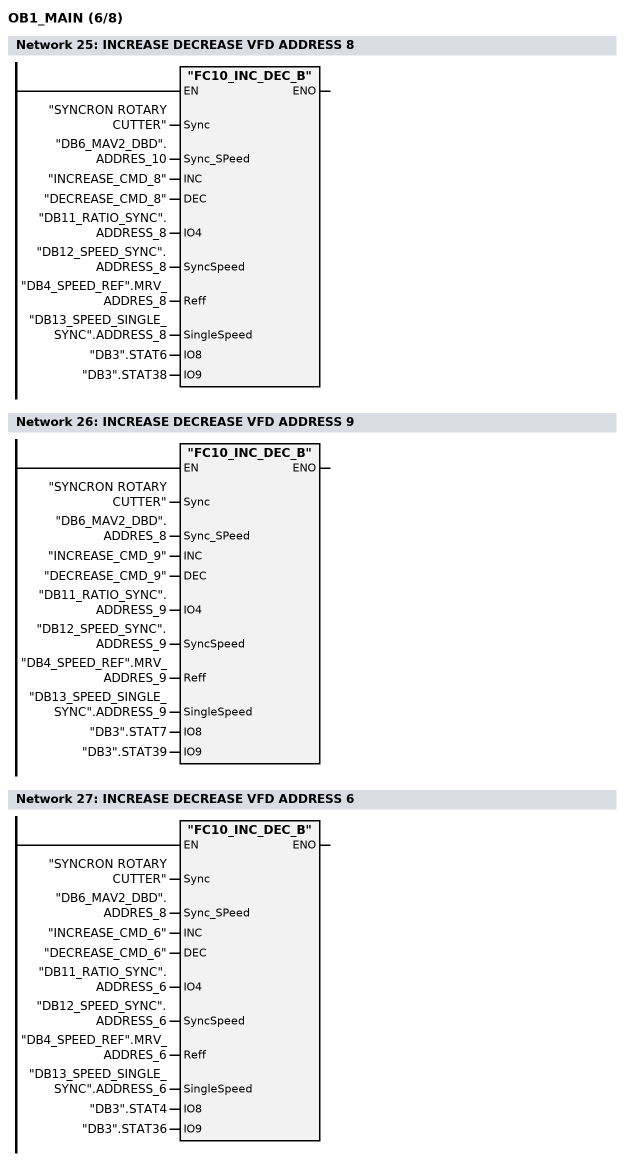
   RUNG wire#powerrail
      "FC10_INC_DEC_B"(Sync := "SYNCRON ROTARY CUTTER", Sync_SPeed := "DB6_MAV2_DBD".ADDRES_10, INC := "INCREASE_CMD_8", DEC := "DECREASE_CMD_8", IO4 := "DB11_RATIO_SYNC".ADDRESS_8, SyncSpeed := "DB12_SPEED_SYNC".ADDRESS_8, Reff := "DB4_SPEED_REF".MRV_ADDRES_8, SingleSpeed := "DB13_SPEED_SINGLE_SYNC".ADDRESS_8, IO8 := "DB3".STAT6, IO9 := "DB3".STAT38)
   END_RUNG
   // the same network as SCL:
   "FC10_INC_DEC_B"(Sync := "SYNCRON ROTARY CUTTER",
                    Sync_SPeed := "DB6_MAV2_DBD".ADDRES_10,
                    INC := "INCREASE_CMD_8",
                    DEC := "DECREASE_CMD_8",
                    IO4 := "DB11_RATIO_SYNC".ADDRESS_8,
                    SyncSpeed := "DB12_SPEED_SYNC".ADDRESS_8,
                    Reff := "DB4_SPEED_REF".MRV_ADDRES_8,
                    SingleSpeed := "DB13_SPEED_SINGLE_SYNC".ADDRESS_8,
                    IO8 := "DB3".STAT6,
                    IO9 := "DB3".STAT38);
END_REGION

REGION Network 26: INCREASE DECREASE VFD ADDRESS 9
   RUNG wire#powerrail
      "FC10_INC_DEC_B"(Sync := "SYNCRON ROTARY CUTTER", Sync_SPeed := "DB6_MAV2_DBD".ADDRES_8, INC := "INCREASE_CMD_9", DEC := "DECREASE_CMD_9", IO4 := "DB11_RATIO_SYNC".ADDRESS_9, SyncSpeed := "DB12_SPEED_SYNC".ADDRESS_9, Reff := "DB4_SPEED_REF".MRV_ADDRES_9, SingleSpeed := "DB13_SPEED_SINGLE_SYNC".ADDRESS_9, IO8 := "DB3".STAT7, IO9 := "DB3".STAT39)
   END_RUNG
   // the same network as SCL:
   "FC10_INC_DEC_B"(Sync := "SYNCRON ROTARY CUTTER",
                    Sync_SPeed := "DB6_MAV2_DBD".ADDRES_8,
                    INC := "INCREASE_CMD_9",
                    DEC := "DECREASE_CMD_9",
                    IO4 := "DB11_RATIO_SYNC".ADDRESS_9,
                    SyncSpeed := "DB12_SPEED_SYNC".ADDRESS_9,
                    Reff := "DB4_SPEED_REF".MRV_ADDRES_9,
                    SingleSpeed := "DB13_SPEED_SINGLE_SYNC".ADDRESS_9,
                    IO8 := "DB3".STAT7,
                    IO9 := "DB3".STAT39);
END_REGION

REGION Network 27: INCREASE DECREASE VFD ADDRESS 6
   RUNG wire#powerrail
      "FC10_INC_DEC_B"(Sync := "SYNCRON ROTARY CUTTER", Sync_SPeed := "DB6_MAV2_DBD".ADDRES_8, INC := "INCREASE_CMD_6", DEC := "DECREASE_CMD_6", IO4 := "DB11_RATIO_SYNC".ADDRESS_6, SyncSpeed := "DB12_SPEED_SYNC".ADDRESS_6, Reff := "DB4_SPEED_REF".MRV_ADDRES_6, SingleSpeed := "DB13_SPEED_SINGLE_SYNC".ADDRESS_6, IO8 := "DB3".STAT4, IO9 := "DB3".STAT36)
   END_RUNG
   // the same network as SCL:
   "FC10_INC_DEC_B"(Sync := "SYNCRON ROTARY CUTTER",
                    Sync_SPeed := "DB6_MAV2_DBD".ADDRES_8,
                    INC := "INCREASE_CMD_6",
                    DEC := "DECREASE_CMD_6",
                    IO4 := "DB11_RATIO_SYNC".ADDRESS_6,
                    SyncSpeed := "DB12_SPEED_SYNC".ADDRESS_6,
                    Reff := "DB4_SPEED_REF".MRV_ADDRES_6,
                    SingleSpeed := "DB13_SPEED_SINGLE_SYNC".ADDRESS_6,
                    IO8 := "DB3".STAT4,
                    IO9 := "DB3".STAT36);
END_REGION

REGION Network 28: INCREASE DECREASE VFD ADDRESS 7
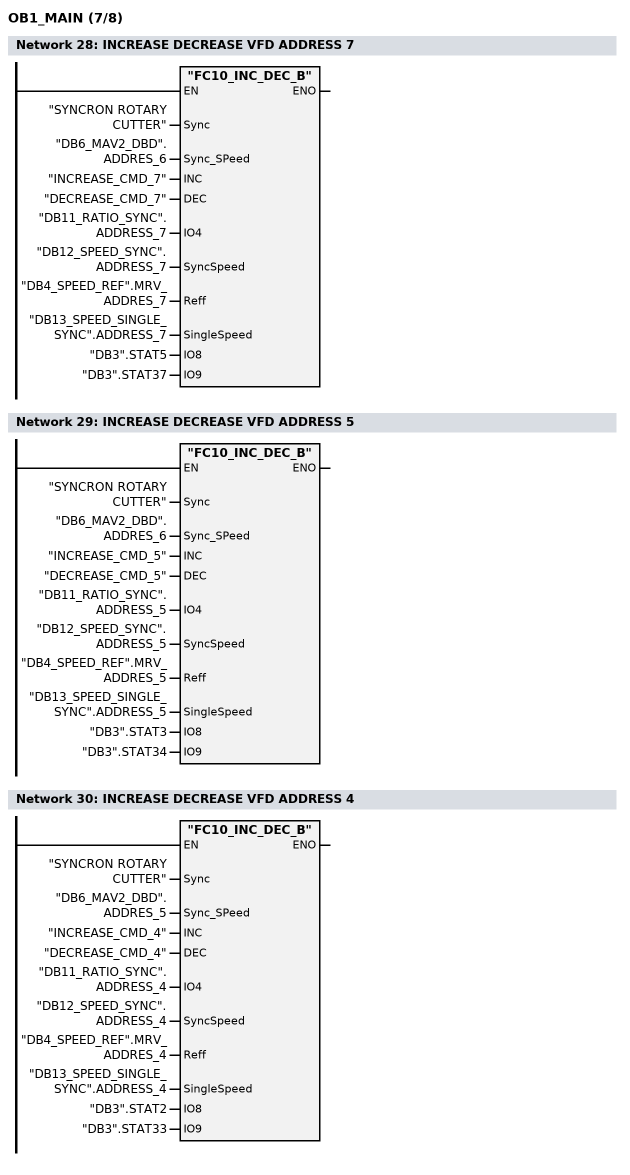
   RUNG wire#powerrail
      "FC10_INC_DEC_B"(Sync := "SYNCRON ROTARY CUTTER", Sync_SPeed := "DB6_MAV2_DBD".ADDRES_6, INC := "INCREASE_CMD_7", DEC := "DECREASE_CMD_7", IO4 := "DB11_RATIO_SYNC".ADDRESS_7, SyncSpeed := "DB12_SPEED_SYNC".ADDRESS_7, Reff := "DB4_SPEED_REF".MRV_ADDRES_7, SingleSpeed := "DB13_SPEED_SINGLE_SYNC".ADDRESS_7, IO8 := "DB3".STAT5, IO9 := "DB3".STAT37)
   END_RUNG
   // the same network as SCL:
   "FC10_INC_DEC_B"(Sync := "SYNCRON ROTARY CUTTER",
                    Sync_SPeed := "DB6_MAV2_DBD".ADDRES_6,
                    INC := "INCREASE_CMD_7",
                    DEC := "DECREASE_CMD_7",
                    IO4 := "DB11_RATIO_SYNC".ADDRESS_7,
                    SyncSpeed := "DB12_SPEED_SYNC".ADDRESS_7,
                    Reff := "DB4_SPEED_REF".MRV_ADDRES_7,
                    SingleSpeed := "DB13_SPEED_SINGLE_SYNC".ADDRESS_7,
                    IO8 := "DB3".STAT5,
                    IO9 := "DB3".STAT37);
END_REGION

REGION Network 29: INCREASE DECREASE VFD ADDRESS 5
   RUNG wire#powerrail
      "FC10_INC_DEC_B"(Sync := "SYNCRON ROTARY CUTTER", Sync_SPeed := "DB6_MAV2_DBD".ADDRES_6, INC := "INCREASE_CMD_5", DEC := "DECREASE_CMD_5", IO4 := "DB11_RATIO_SYNC".ADDRESS_5, SyncSpeed := "DB12_SPEED_SYNC".ADDRESS_5, Reff := "DB4_SPEED_REF".MRV_ADDRES_5, SingleSpeed := "DB13_SPEED_SINGLE_SYNC".ADDRESS_5, IO8 := "DB3".STAT3, IO9 := "DB3".STAT34)
   END_RUNG
   // the same network as SCL:
   "FC10_INC_DEC_B"(Sync := "SYNCRON ROTARY CUTTER",
                    Sync_SPeed := "DB6_MAV2_DBD".ADDRES_6,
                    INC := "INCREASE_CMD_5",
                    DEC := "DECREASE_CMD_5",
                    IO4 := "DB11_RATIO_SYNC".ADDRESS_5,
                    SyncSpeed := "DB12_SPEED_SYNC".ADDRESS_5,
                    Reff := "DB4_SPEED_REF".MRV_ADDRES_5,
                    SingleSpeed := "DB13_SPEED_SINGLE_SYNC".ADDRESS_5,
                    IO8 := "DB3".STAT3,
                    IO9 := "DB3".STAT34);
END_REGION

REGION Network 30: INCREASE DECREASE VFD ADDRESS 4
   RUNG wire#powerrail
      "FC10_INC_DEC_B"(Sync := "SYNCRON ROTARY CUTTER", Sync_SPeed := "DB6_MAV2_DBD".ADDRES_5, INC := "INCREASE_CMD_4", DEC := "DECREASE_CMD_4", IO4 := "DB11_RATIO_SYNC".ADDRESS_4, SyncSpeed := "DB12_SPEED_SYNC".ADDRESS_4, Reff := "DB4_SPEED_REF".MRV_ADDRES_4, SingleSpeed := "DB13_SPEED_SINGLE_SYNC".ADDRESS_4, IO8 := "DB3".STAT2, IO9 := "DB3".STAT33)
   END_RUNG
   // the same network as SCL:
   "FC10_INC_DEC_B"(Sync := "SYNCRON ROTARY CUTTER",
                    Sync_SPeed := "DB6_MAV2_DBD".ADDRES_5,
                    INC := "INCREASE_CMD_4",
                    DEC := "DECREASE_CMD_4",
                    IO4 := "DB11_RATIO_SYNC".ADDRESS_4,
                    SyncSpeed := "DB12_SPEED_SYNC".ADDRESS_4,
                    Reff := "DB4_SPEED_REF".MRV_ADDRES_4,
                    SingleSpeed := "DB13_SPEED_SINGLE_SYNC".ADDRESS_4,
                    IO8 := "DB3".STAT2,
                    IO9 := "DB3".STAT33);
END_REGION

REGION Network 31: INCREASE DECREASE VFD ADDRESS 3
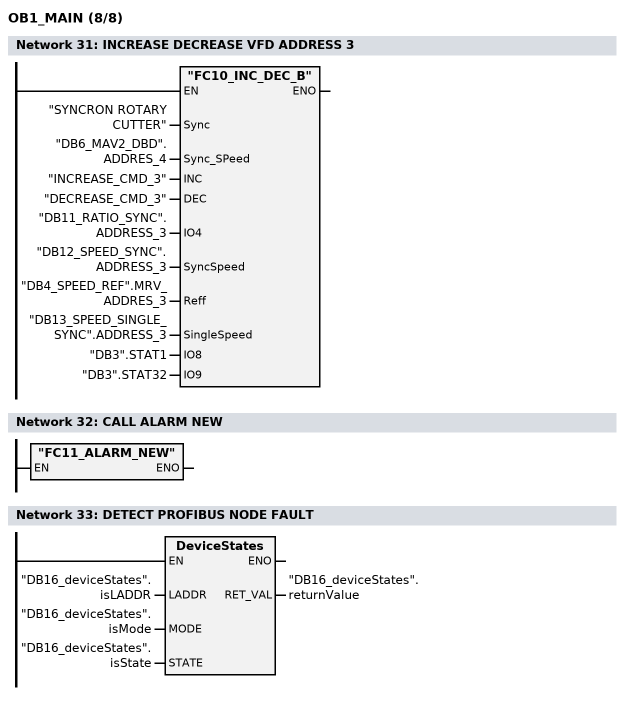
   RUNG wire#powerrail
      "FC10_INC_DEC_B"(Sync := "SYNCRON ROTARY CUTTER", Sync_SPeed := "DB6_MAV2_DBD".ADDRES_4, INC := "INCREASE_CMD_3", DEC := "DECREASE_CMD_3", IO4 := "DB11_RATIO_SYNC".ADDRESS_3, SyncSpeed := "DB12_SPEED_SYNC".ADDRESS_3, Reff := "DB4_SPEED_REF".MRV_ADDRES_3, SingleSpeed := "DB13_SPEED_SINGLE_SYNC".ADDRESS_3, IO8 := "DB3".STAT1, IO9 := "DB3".STAT32)
   END_RUNG
   // the same network as SCL:
   "FC10_INC_DEC_B"(Sync := "SYNCRON ROTARY CUTTER",
                    Sync_SPeed := "DB6_MAV2_DBD".ADDRES_4,
                    INC := "INCREASE_CMD_3",
                    DEC := "DECREASE_CMD_3",
                    IO4 := "DB11_RATIO_SYNC".ADDRESS_3,
                    SyncSpeed := "DB12_SPEED_SYNC".ADDRESS_3,
                    Reff := "DB4_SPEED_REF".MRV_ADDRES_3,
                    SingleSpeed := "DB13_SPEED_SINGLE_SYNC".ADDRESS_3,
                    IO8 := "DB3".STAT1,
                    IO9 := "DB3".STAT32);
END_REGION

REGION Network 32: CALL ALARM NEW
   RUNG wire#powerrail
      "FC11_ALARM_NEW"()
   END_RUNG
   // the same network as SCL:
   "FC11_ALARM_NEW"();
END_REGION

REGION Network 33: DETECT PROFIBUS NODE FAULT
   // no SCL statement known for DeviceStates: written as a call
   "DB16_deviceStates".returnValue := DeviceStates(LADDR := "DB16_deviceStates".isLADDR,
                           MODE := "DB16_deviceStates".isMode,
                           STATE := "DB16_deviceStates".isState);
END_REGION
END_ORGANIZATION_BLOCK

ORGANIZATION_BLOCK "OB80_TIME_ERROR"   // OB80, LAD, TimeErrorInterrupt
{ S7_Optimized_Access := 'FALSE' }
VERSION : 0.1
   VAR_TEMP
      TEMP0 : Byte;
      TEMP1 : Byte;
      TEMP2 : Byte;
      TEMP3 : Byte;
      TEMP4 : Byte;
      TEMP5 : Byte;
      TEMP6 : Word;
      TEMP7 : Byte;
      TEMP8 : Byte;
      TEMP9 : Byte;
      TEMP10 : Byte;
      TEMP11 : Date_And_Time;
   END_VAR
BEGIN
END_ORGANIZATION_BLOCK

ORGANIZATION_BLOCK "OB82_DIAG_INTERRUPT"   // OB82, LAD, DiagnosticErrorInterrupt
{ S7_Optimized_Access := 'FALSE' }
VERSION : 0.1
   VAR_TEMP
      TEMP0 : Byte;
      TEMP1 : Byte;
      TEMP2 : Byte;
      TEMP3 : Byte;
      TEMP4 : Byte;
      TEMP5 : Byte;
      TEMP6 : Word;
      TEMP7 : Byte;
      TEMP8 : Byte;
      TEMP9 : Byte;
      TEMP10 : Byte;
      TEMP11 : Date_And_Time;
   END_VAR
BEGIN
END_ORGANIZATION_BLOCK

ORGANIZATION_BLOCK "OB83_Pull or plug of modules"   // OB83, LAD, PullPlug
{ S7_Optimized_Access := 'TRUE' }
VERSION : 0.1
   VAR_INPUT
      LADDR : Hw_Io;   // Hardware identifier
      Event_Class : Byte;   // 16#38/39: module inserted, removed
      Fault_ID : Byte;   // Fault identifier
   END_VAR
BEGIN
END_ORGANIZATION_BLOCK

ORGANIZATION_BLOCK "OB86_RACK_FAILURE"   // OB86, LAD, RackStationFailure
{ S7_Optimized_Access := 'FALSE' }
VERSION : 0.1
   VAR_TEMP
      TEMP0 : Byte;
      TEMP1 : Byte;
      TEMP2 : Byte;
      TEMP3 : Byte;
      TEMP4 : Byte;
      TEMP5 : Byte;
      TEMP6 : Word;
      TEMP7 : Byte;
      TEMP8 : Byte;
      TEMP9 : Byte;
      TEMP10 : Byte;
      TEMP11 : Date_And_Time;
   END_VAR
BEGIN
END_ORGANIZATION_BLOCK

ORGANIZATION_BLOCK "OB100_STARTUP_MODE"   // OB100, LAD, Startup
{ S7_Optimized_Access := 'FALSE' }
VERSION : 0.1
   VAR_TEMP
      TEMP0 : Byte;
      TEMP1 : Byte;
      TEMP2 : Byte;
      TEMP3 : Byte;
      TEMP4 : Byte;
      TEMP5 : Byte;
      TEMP6 : Word;
      TEMP7 : Byte;
      TEMP8 : Byte;
      TEMP9 : Byte;
      TEMP10 : Byte;
      TEMP11 : Date_And_Time;
   END_VAR
BEGIN
END_ORGANIZATION_BLOCK

ORGANIZATION_BLOCK "OB121_PROGRAMMING_ERR"   // OB121, LAD, ProgrammingError
{ S7_Optimized_Access := 'FALSE' }
VERSION : 0.1
   VAR_TEMP
      TEMP0 : Byte;
      TEMP1 : Byte;
      TEMP2 : Byte;
      TEMP3 : Byte;
      TEMP4 : Byte;
      TEMP5 : Byte;
      TEMP6 : Word;
      TEMP7 : Byte;
      TEMP8 : Byte;
      TEMP9 : Byte;
      TEMP10 : Byte;
      TEMP11 : Date_And_Time;
   END_VAR
BEGIN
END_ORGANIZATION_BLOCK

ORGANIZATION_BLOCK "OB122_I/O_ACCES_ERR"   // OB122, LAD, IOAccessError
{ S7_Optimized_Access := 'FALSE' }
VERSION : 0.1
   VAR_TEMP
      TEMP0 : Byte;
      TEMP1 : Byte;
      TEMP2 : Byte;
      TEMP3 : Byte;
      TEMP4 : Byte;
      TEMP5 : Byte;
      TEMP6 : Word;
      TEMP7 : Byte;
      TEMP8 : Byte;
      TEMP9 : Byte;
      TEMP10 : Byte;
      TEMP11 : Date_And_Time;
   END_VAR
BEGIN
END_ORGANIZATION_BLOCK

(* ===== HMI "HMI_RT_1" =====
system functions are stored by id; their names below are inferred from use
connection "SPS_1": ETHERNET, SMART_S7_1500_OMS

HMI tags "Default tag table"
   "Tag_ScreenNumber" : UInt, internal

HMI tags "Animation_control"
   "animation_page" : Int, internal

HMI tags "Speed Reference"
   "speedReff_singleSync_address_2" : Real AT %DB13.DBD8, 1 s
   "speedReff_singleSync_address_3" : Real AT %DB13.DBD12, 1 s
   "speedReff_singleSync_address_4" : Real AT %DB13.DBD16, 1 s
   "speedReff_singleSync_address_5" : Real AT %DB13.DBD20, 1 s
   "speedReff_singleSync_address_6" : Real AT %DB13.DBD24, 1 s
   "speedReff_singleSync_address_7" : Real AT %DB13.DBD28, 1 s
   "speedReff_singleSync_address_8" : Real AT %DB13.DBD32, 1 s
   "speedReff_singleSync_address_9" : Real AT %DB13.DBD36, 1 s
   "speedReff_singleSync_address_10" : Real AT %DB13.DBD40, 1 s
   "speedReff_singleSync_address_11" : Real AT %DB13.DBD44, 1 s
   "speedReff_singleSync_address_12" : Real AT %DB13.DBD48, 1 s
   "speedReff_singleSync_address_13" : Real AT %DB13.DBD52, 1 s
   "speedReff_singleSync_address_14" : Real AT %DB13.DBD56, 1 s
   "speedReff_singleSync_address_15" : Real AT %DB13.DBD60, 1 s
   "speedReff_singleSync_address_16" : Real AT %DB13.DBD64, 1 s
   "speedReff_singleSync_address_17" : Real AT %DB13.DBD68, 1 s
   "speedReff_singleSync_address_18" : Real AT %DB13.DBD72, 1 s
   "speedReff_singleSync_address_19" : Real AT %DB13.DBD76, 1 s
   "speedReff_singleSync_address_20" : Real AT %DB13.DBD80, 1 s
   "speedReff_singleSync_address_21" : Real AT %DB13.DBD84, 1 s
   "speedReff_singleSync_address_22" : Real AT %DB13.DBD88, 1 s
   "speedReff_singleSync_address_23" : Real AT %DB13.DBD92, 1 s
   "speedReff_NOT_singleSync_address_3" : Real AT %DB12.DBD4, 1 s
   "speedReff_NOT_singleSync_address_4" : Real AT %DB12.DBD8, 1 s
   "speedReff_NOT_singleSync_address_5" : Real AT %DB12.DBD12, 1 s
   "speedReff_NOT_singleSync_address_6" : Real AT %DB12.DBD16, 1 s
   "speedReff_NOT_singleSync_address_7" : Real AT %DB12.DBD20, 1 s
   "speedReff_NOT_singleSync_address_8" : Real AT %DB12.DBD24, 1 s
   "speedReff_NOT_singleSync_address_9" : Real AT %DB12.DBD28, 1 s
   "speedReff_NOT_singleSync_address_10" : Real AT %DB12.DBD32, 1 s
   "speedReff_NOT_singleSync_address_11" : Real AT %DB12.DBD36, 1 s
   "speedReff_NOT_singleSync_address_12" : Real AT %DB12.DBD40, 1 s
   "speedReff_NOT_singleSync_address_13" : Real AT %DB12.DBD44, 1 s
   "speedReff_NOT_singleSync_address_14" : Real AT %DB12.DBD48, 1 s
   "speedReff_NOT_singleSync_address_15" : Real AT %DB12.DBD52, 1 s
   "speedReff_NOT_singleSync_address_16" : Real AT %DB12.DBD56, 1 s
   "speedReff_NOT_singleSync_address_17" : Real AT %DB12.DBD60, 1 s
   "speedReff_NOT_singleSync_address_18" : Real AT %DB12.DBD64, 1 s
   "speedReff_NOT_singleSync_address_19" : Real AT %DB12.DBD68, 1 s
   "speedReff_NOT_singleSync_address_20" : Real AT %DB12.DBD72, 1 s
   "speedReff_NOT_singleSync_address_21" : Real AT %DB12.DBD76, 1 s
   "speedReff_NOT_singleSync_address_22" : Real AT %DB12.DBD80, 1 s
   "speedReff_NOT_singleSync_address_23" : Real AT %DB12.DBD84, 1 s

HMI tags "Speed Actual"
   "speedActual_address_2" : Real AT %DB6.DBD116, 1 s
   "speedActual_address_3" : Real AT %DB6.DBD120, 1 s
   "speedActual_address_4" : Real AT %DB6.DBD124, 1 s
   "speedActual_address_5" : Real AT %DB6.DBD128, 1 s
   "speedActual_address_6" : Real AT %DB6.DBD132, 1 s
   "speedActual_address_7" : Real AT %DB6.DBD136, 1 s
   "speedActual_address_8" : Real AT %DB6.DBD140, 1 s
   "speedActual_address_9" : Real AT %DB6.DBD144, 1 s
   "speedActual_address_10" : Real AT %DB6.DBD148, 1 s
   "speedActual_address_11" : Real AT %DB6.DBD152, 1 s
   "speedActual_address_12" : Real AT %DB6.DBD156, 1 s
   "speedActual_address_13" : Real AT %DB6.DBD160, 1 s
   "speedActual_address_14" : Real AT %DB6.DBD164, 1 s
   "speedActual_address_15" : Real AT %DB6.DBD168, 1 s
   "speedActual_address_16" : Real AT %DB6.DBD172, 1 s
   "speedActual_address_17" : Real AT %DB6.DBD176, 1 s
   "speedActual_address_18" : Real AT %DB6.DBD180, 1 s
   "speedActual_address_19" : Real AT %DB6.DBD184, 1 s
   "speedActual_address_20" : Real AT %DB6.DBD188, 1 s
   "speedActual_address_21" : Real AT %DB6.DBD192, 1 s
   "speedActual_address_22" : Real AT %DB6.DBD196, 1 s
   "speedActual_address_23" : Real AT %DB6.DBD200, 1 s

HMI tags "Control_Speed"
   "increaseSpeed_address_2" : Bool AT %M20.1, 1 s
   "increaseSpeed_address_3" : Bool AT %M20.2, 1 s
   "increaseSpeed_address_4" : Bool AT %M20.3, 1 s
   "increaseSpeed_address_5" : Bool AT %M20.4, 1 s
   "increaseSpeed_address_6" : Bool AT %M20.5, 1 s
   "increaseSpeed_address_7" : Bool AT %M20.6, 1 s
   "increaseSpeed_address_8" : Bool AT %M20.7, 1 s
   "increaseSpeed_address_9" : Bool AT %M21.0, 1 s
   "increaseSpeed_address_10" : Bool AT %M21.1, 1 s
   "increaseSpeed_address_11" : Bool AT %M21.2, 1 s
   "increaseSpeed_address_12" : Bool AT %M21.3, 1 s
   "increaseSpeed_address_13" : Bool AT %M21.4, 1 s
   "increaseSpeed_address_14" : Bool AT %M21.5, 1 s
   "increaseSpeed_address_15" : Bool AT %M21.6, 1 s
   "increaseSpeed_address_16" : Bool AT %M21.7, 1 s
   "increaseSpeed_address_17" : Bool AT %M22.0, 1 s
   "increaseSpeed_address_18" : Bool AT %M22.1, 1 s
   "increaseSpeed_address_19" : Bool AT %M22.2, 1 s
   "increaseSpeed_address_20" : Bool AT %M22.3, 1 s
   "increaseSpeed_address_21" : Bool AT %M22.4, 1 s
   "increaseSpeed_address_22" : Bool AT %M22.5, 1 s
   "increaseSpeed_address_23" : Bool AT %M22.6, 1 s
   "decreaseSpeed_address_2" : Bool AT %M24.1, 1 s
   "decreaseSpeed_address_3" : Bool AT %M24.2, 1 s
   "decreaseSpeed_address_4" : Bool AT %M24.3, 1 s
   "decreaseSpeed_address_5" : Bool AT %M24.4, 1 s
   "decreaseSpeed_address_6" : Bool AT %M24.5, 1 s
   "decreaseSpeed_address_7" : Bool AT %M24.6, 1 s
   "decreaseSpeed_address_8" : Bool AT %M24.7, 1 s
   "decreaseSpeed_address_9" : Bool AT %M25.0, 1 s
   "decreaseSpeed_address_10" : Bool AT %M25.1, 1 s
   "decreaseSpeed_address_11" : Bool AT %M25.2, 1 s
   "decreaseSpeed_address_12" : Bool AT %M25.3, 1 s
   "decreaseSpeed_address_13" : Bool AT %M25.4, 1 s
   "decreaseSpeed_address_14" : Bool AT %M25.5, 1 s
   "decreaseSpeed_address_15" : Bool AT %M25.6, 1 s
   "decreaseSpeed_address_16" : Bool AT %M25.7, 1 s
   "decreaseSpeed_address_17" : Bool AT %M26.0, 1 s
   "decreaseSpeed_address_18" : Bool AT %M26.1, 1 s
   "decreaseSpeed_address_19" : Bool AT %M26.2, 1 s
   "decreaseSpeed_address_20" : Bool AT %M26.3, 1 s
   "decreaseSpeed_address_21" : Bool AT %M26.4, 1 s
   "decreaseSpeed_address_22" : Bool AT %M26.5, 1 s
   "decreaseSpeed_address_23" : Bool AT %M26.6, 1 s
   "statusIncrease_address_2" : Bool AT %M10.0, 1 s
   "statusIncrease_address_3" : Bool AT %M10.1, 1 s
   "statusIncrease_address_4" : Bool AT %M10.2, 1 s
   "statusIncrease_address_5" : Bool AT %M10.3, 1 s
   "statusIncrease_address_6" : Bool AT %M10.4, 1 s
   "statusIncrease_address_7" : Bool AT %M10.5, 1 s
   "statusIncrease_address_8" : Bool AT %M10.6, 1 s
   "statusIncrease_address_9" : Bool AT %M10.7, 1 s
   "statusIncrease_address_10" : Bool AT %M11.0, 1 s
   "statusIncrease_address_11" : Bool AT %M11.1, 1 s
   "statusIncrease_address_12" : Bool AT %M11.2, 1 s
   "statusIncrease_address_13" : Bool AT %M11.3, 1 s
   "statusIncrease_address_14" : Bool AT %M11.4, 1 s
   "statusIncrease_address_15" : Bool AT %M11.5, 1 s
   "statusIncrease_address_16" : Bool AT %M11.6, 1 s
   "statusIncrease_address_17" : Bool AT %M11.7, 1 s
   "statusIncrease_address_18" : Bool AT %M12.0, 1 s
   "statusIncrease_address_19" : Bool AT %M12.1, 1 s
   "statusIncrease_address_20" : Bool AT %M12.2, 1 s
   "statusIncrease_address_21" : Bool AT %M12.3, 1 s
   "statusIncrease_address_22" : Bool AT %M12.4, 1 s
   "statusIncrease_address_23" : Bool AT %M12.5, 1 s
   "statusDecrease_address_2" : Bool AT %M15.1, 1 s
   "statusDecrease_address_3" : Bool AT %M15.2, 1 s
   "statusDecrease_address_4" : Bool AT %M15.3, 1 s
   "statusDecrease_address_5" : Bool AT %M15.4, 1 s
   "statusDecrease_address_6" : Bool AT %M15.5, 1 s
   "statusDecrease_address_7" : Bool AT %M15.6, 1 s
   "statusDecrease_address_8" : Bool AT %M15.7, 1 s
   "statusDecrease_address_9" : Bool AT %M16.0, 1 s
   "statusDecrease_address_10" : Bool AT %M16.1, 1 s
   "statusDecrease_address_11" : Bool AT %M16.2, 1 s
   "statusDecrease_address_12" : Bool AT %M16.3, 1 s
   "statusDecrease_address_13" : Bool AT %M16.4, 1 s
   "statusDecrease_address_14" : Bool AT %M16.5, 1 s
   "statusDecrease_address_15" : Bool AT %M16.6, 1 s
   "statusDecrease_address_16" : Bool AT %M16.7, 1 s
   "statusDecrease_address_17" : Bool AT %M17.0, 1 s
   "statusDecrease_address_18" : Bool AT %M17.1, 1 s
   "statusDecrease_address_19" : Bool AT %M17.2, 1 s
   "statusDecrease_address_20" : Bool AT %M17.3, 1 s
   "statusDecrease_address_21" : Bool AT %M17.4, 1 s
   "statusDecrease_address_22" : Bool AT %M17.5, 1 s
   "statusDecrease_address_23" : Bool AT %M17.6, 1 s

HMI tags "Mode"
   "Syncron_1" : Bool AT %I6.5, 1 s
   "Syncron_2" : Bool AT %I6.6, 1 s
   "Syncron_3" : Bool AT %I6.7, 1 s
   "Rotary_Cutting" : Bool AT %I7.1, 1 s
   "Rotary_Moulder" : Bool AT %I7.0, 1 s

HMI tags "Alarm"
   "Alarm_Adress_2" : Word AT %DB15.DBW0, 1 s
   "Alarm_Adress_3" : Word AT %DB15.DBW2, 1 s
   "Alarm_Adress_4" : Word AT %DB15.DBW4, 1 s
   "Alarm_Adress_5" : Word AT %DB15.DBW6, 1 s
   "Alarm_Adress_6" : Word AT %DB15.DBW8, 1 s
   "Alarm_Adress_7" : Word AT %DB15.DBW10, 1 s
   "Alarm_Adress_8" : Word AT %DB15.DBW12, 1 s
   "Alarm_Adress_9" : Word AT %DB15.DBW14, 1 s
   "Alarm_Adress_10" : Word AT %DB15.DBW16, 1 s
   "Alarm_Adress_11" : Word AT %DB15.DBW18, 1 s
   "Alarm_Adress_12" : Word AT %DB15.DBW20, 1 s
   "Alarm_Adress_13" : Word AT %DB15.DBW22, 1 s
   "Alarm_Adress_14" : Word AT %DB15.DBW24, 1 s
   "Alarm_Adress_15" : Word AT %DB15.DBW26, 1 s
   "Alarm_Adress_16" : Word AT %DB15.DBW28, 1 s
   "Alarm_Adress_17" : Word AT %DB15.DBW30, 1 s
   "Alarm_Adress_18" : Word AT %DB15.DBW32, 1 s
   "Alarm_Adress_19" : Word AT %DB15.DBW34, 1 s
   "Alarm_Adress_20" : Word AT %DB15.DBW36, 1 s
   "Alarm_Adress_21" : Word AT %DB15.DBW38, 1 s
   "Alarm_Adress_22" : Word AT %DB15.DBW40, 1 s
   "Alarm_Adress_23" : Word AT %DB15.DBW42, 1 s
   "EMERGENCY" : Bool AT %M92.7, 1 s

HMI tags "Profibus_Status"
   "Address_2" : Bool AT %M90.1, 1 s
   "Address_3" : Bool AT %M90.2, 1 s
   "Address_4" : Bool AT %M90.3, 1 s
   "Address_5" : Bool AT %M90.4, 1 s
   "Address_6" : Bool AT %M90.5, 1 s
   "Address_7" : Bool AT %M90.6, 1 s
   "Address_8" : Bool AT %M90.7, 1 s
   "Address_9" : Bool AT %M91.0, 1 s
   "Address_10" : Bool AT %M91.1, 1 s
   "Address_11" : Bool AT %M91.2, 1 s
   "Address_12" : Bool AT %M91.3, 1 s
   "Address_13" : Bool AT %M91.4, 1 s
   "Address_14" : Bool AT %M91.5, 1 s
   "Address_15" : Bool AT %M91.6, 1 s
   "Address_16" : Bool AT %M91.7, 1 s
   "Address_17" : Bool AT %M92.0, 1 s
   "Address_18" : Bool AT %M92.1, 1 s
   "Address_19" : Bool AT %M92.2, 1 s
   "Address_20" : Bool AT %M92.3, 1 s
   "Address_21" : Bool AT %M92.4, 1 s
   "Address_22" : Bool AT %M92.5, 1 s
   "Address_23" : Bool AT %M92.6, 1 s
   "Alarm_1" : Word AT %MW90, 1 s
   "Alarm_2" : Word AT %MW92, 1 s

HMI tags "Motor Running Status"
   "Running_Motor Addres_2" : Bool AT %DB15.DBX0.3, 1 s
   "Running_Motor Addres_3" : Bool AT %DB15.DBX2.3, 1 s
   "Running_Motor Addres_4" : Bool AT %DB15.DBX4.3, 1 s
   "Running_Motor Addres_5" : Bool AT %DB15.DBX6.3, 1 s
   "Running_Motor Addres_6" : Bool AT %DB15.DBX8.3, 1 s
   "Running_Motor Addres_7" : Bool AT %DB15.DBX10.3, 1 s
   "Running_Motor Addres_8" : Bool AT %DB15.DBX12.3, 1 s
   "Running_Motor Addres_9" : Bool AT %DB15.DBX14.3, 1 s
   "Running_Motor Addres_10" : Bool AT %DB15.DBX16.3, 1 s
   "Running_Motor Addres_11" : Bool AT %DB15.DBX18.3, 1 s
   "Running_Motor Addres_12" : Bool AT %DB15.DBX20.3, 1 s
   "Running_Motor Addres_13" : Bool AT %DB15.DBX22.3, 1 s
   "Running_Motor Addres_14" : Bool AT %DB15.DBX24.3, 1 s
   "Running_Motor Addres_15" : Bool AT %DB15.DBX26.3, 1 s
   "Running_Motor Addres_16" : Bool AT %DB15.DBX28.3, 1 s
   "Running_Motor Addres_17" : Bool AT %DB15.DBX30.3, 1 s
   "Running_Motor Addres_18" : Bool AT %DB15.DBX32.3, 1 s
   "Running_Motor Addres_19" : Bool AT %DB15.DBX34.3, 1 s
   "Running_Motor Addres_20" : Bool AT %DB15.DBX36.3, 1 s
   "Running_Motor Addres_21" : Bool AT %DB15.DBX38.3, 1 s
   "Running_Motor Addres_22" : Bool AT %DB15.DBX40.3, 1 s
   "Running_Motor Addres_23" : Bool AT %DB15.DBX42.3, 1 s

HMI tags "DI/DO"
   "In_125_0" : Bool AT %I125.0, 1 s
   "In_125_1" : Bool AT %I125.1, 1 s
   "In_125_2" : Bool AT %I125.2, 1 s
   "In_125_3" : Bool AT %I125.3, 1 s
   "In_125_4" : Bool AT %I125.4, 1 s
   "In_125_5" : Bool AT %I125.5, 1 s
   "In_125_6" : Bool AT %I125.6, 1 s
   "In_125_7" : Bool AT %I125.7, 1 s
   "In_124_0" : Bool AT %I124.0, 1 s
   "In_124_1" : Bool AT %I124.1, 1 s
   "In_124_2" : Bool AT %I124.2, 1 s
   "In_124_3" : Bool AT %I124.3, 1 s
   "In_124_4" : Bool AT %I124.4, 1 s
   "In_124_5" : Bool AT %I124.5, 1 s
   "In_124_6" : Bool AT %I124.6, 1 s
   "In_124_7" : Bool AT %I124.7, 1 s
   "In_126_0" : Bool AT %I126.0, 1 s
   "In_126_1" : Bool AT %I126.1, 1 s
   "In_126_2" : Bool AT %I126.2, 1 s
   "In_126_3" : Bool AT %I126.3, 1 s
   "In_126_4" : Bool AT %I126.4, 1 s
   "In_126_5" : Bool AT %I126.5, 1 s
   "In_126_6" : Bool AT %I126.6, 1 s
   "In_126_7" : Bool AT %I126.7, 1 s
   "In_127_0" : Bool AT %I127.0, 1 s
   "In_127_1" : Bool AT %I127.1, 1 s
   "In_127_2" : Bool AT %I127.2, 1 s
   "In_127_3" : Bool AT %I127.3, 1 s
   "In_127_4" : Bool AT %I127.4, 1 s
   "In_127_5" : Bool AT %I127.5, 1 s
   "In_127_6" : Bool AT %I127.6, 1 s
   "In_127_7" : Bool AT %I127.7, 1 s
   "In_0_0" : Bool AT %I0.0, 1 s
   "In_0_1" : Bool AT %I0.1, 1 s
   "In_0_2" : Bool AT %I0.2, 1 s
   "In_0_3" : Bool AT %I0.3, 1 s
   "In_0_4" : Bool AT %I0.4, 1 s
   "In_0_5" : Bool AT %I0.5, 1 s
   "In_0_6" : Bool AT %I0.6, 1 s
   "In_0_7" : Bool AT %I0.7, 1 s
   "In_1_0" : Bool AT %I1.0, 1 s
   "In_1_1" : Bool AT %I1.1, 1 s
   "In_1_2" : Bool AT %I1.2, 1 s
   "In_1_3" : Bool AT %I1.3, 1 s
   "In_1_4" : Bool AT %I1.4, 1 s
   "In_1_5" : Bool AT %I1.5, 1 s
   "In_1_6" : Bool AT %I1.6, 1 s
   "In_1_7" : Bool AT %I1.7, 1 s
   "In_2_0" : Bool AT %I2.0, 1 s
   "In_2_1" : Bool AT %I2.1, 1 s
   "In_2_2" : Bool AT %I2.2, 1 s
   "In_2_3" : Bool AT %I2.3, 1 s
   "In_2_4" : Bool AT %I2.4, 1 s
   "In_2_5" : Bool AT %I2.5, 1 s
   "In_2_6" : Bool AT %I2.6, 1 s
   "In_2_7" : Bool AT %I2.7, 1 s
   "In_3_0" : Bool AT %I3.0, 1 s
   "In_3_1" : Bool AT %I3.1, 1 s
   "In_3_2" : Bool AT %I3.2, 1 s
   "In_3_3" : Bool AT %I3.3, 1 s
   "In_3_4" : Bool AT %I3.4, 1 s
   "In_3_5" : Bool AT %I3.5, 1 s
   "In_3_6" : Bool AT %I3.6, 1 s
   "In_3_7" : Bool AT %I3.7, 1 s
   "In_4_0" : Bool AT %I4.0, 1 s
   "In_4_1" : Bool AT %I4.1, 1 s
   "In_4_2" : Bool AT %I4.2, 1 s
   "In_4_3" : Bool AT %I4.3, 1 s
   "In_4_4" : Bool AT %I4.4, 1 s
   "In_4_5" : Bool AT %I4.5, 1 s
   "In_4_6" : Bool AT %I4.6, 1 s
   "In_4_7" : Bool AT %I4.7, 1 s
   "In_5_0" : Bool AT %I5.0, 1 s
   "In_5_1" : Bool AT %I5.1, 1 s
   "In_5_2" : Bool AT %I5.2, 1 s
   "In_5_3" : Bool AT %I5.3, 1 s
   "In_5_4" : Bool AT %I5.4, 1 s
   "In_5_5" : Bool AT %I5.5, 1 s
   "In_5_6" : Bool AT %I5.6, 1 s
   "In_5_7" : Bool AT %I5.7, 1 s
   "In_6_0" : Bool AT %I6.0, 1 s
   "In_6_1" : Bool AT %I6.1, 1 s
   "In_6_2" : Bool AT %I6.2, 1 s
   "In_6_3" : Bool AT %I6.3, 1 s
   "In_6_4" : Bool AT %I6.4, 1 s
   "In_6_5" : Bool AT %I6.5, 1 s
   "In_6_6" : Bool AT %I6.6, 1 s
   "In_6_7" : Bool AT %I6.7, 1 s
   "In_7_0" : Bool AT %I7.0, 1 s
   "In_7_1" : Bool AT %I7.1, 1 s
   "In_7_2" : Bool AT %I7.2, 1 s
   "In_7_3" : Bool AT %I7.3, 1 s
   "In_7_4" : Bool AT %I7.4, 1 s
   "In_7_5" : Bool AT %I7.5, 1 s
   "In_7_6" : Bool AT %I7.6, 1 s
   "In_7_7" : Bool AT %I7.7, 1 s
   "Out_124_0" : Bool AT %Q124.0, 1 s
   "Out_124_1" : Bool AT %Q124.1, 1 s
   "Out_124_2" : Bool AT %Q124.2, 1 s
   "Out_124_3" : Bool AT %Q124.3, 1 s
   "Out_124_4" : Bool AT %Q124.4, 1 s
   "Out_124_5" : Bool AT %Q124.5, 1 s
   "Out_124_6" : Bool AT %Q124.6, 1 s
   "Out_124_7" : Bool AT %Q124.7, 1 s
   "Out_125_0" : Bool AT %Q125.0, 1 s
   "Out_125_1" : Bool AT %Q125.1, 1 s
   "Out_125_2" : Bool AT %Q125.2, 1 s
   "Out_125_3" : Bool AT %Q125.3, 1 s
   "Out_125_4" : Bool AT %Q125.4, 1 s
   "Out_125_5" : Bool AT %Q125.5, 1 s
   "Out_125_6" : Bool AT %Q125.6, 1 s
   "Out_125_7" : Bool AT %Q125.7, 1 s

discrete alarms
   1: 'Motor 2 Trip', class Errors, trigger "Alarm_Adress_2" bit 3
   2: 'Motor 2 Warning', class Warnings, trigger "Alarm_Adress_2" bit 7
   3: 'Motor 2 Voltage Fault', class Errors, trigger "Alarm_Adress_2" bit 13
   4: 'Motor 2 Torque Fault', class Errors, trigger "Alarm_Adress_2" bit 14
   5: 'Motor 2 Thermal Warning', class Warnings, trigger "Alarm_Adress_2" bit 15
   6: 'Motor 3 Trip', class Errors, trigger "Alarm_Adress_3" bit 3
   7: 'Motor 3 Warning', class Warnings, trigger "Alarm_Adress_3" bit 7
   8: 'Motor 3 Voltage Fault', class Errors, trigger "Alarm_Adress_3" bit 13
   9: 'Motor 3 Torque Fault', class Errors, trigger "Alarm_Adress_3" bit 14
   10: 'Motor 3 Thermal Warning', class Warnings, trigger "Alarm_Adress_3" bit 15
   11: 'Motor 4 Trip', class Errors, trigger "Alarm_Adress_4" bit 3
   12: 'Motor 4 Warning', class Warnings, trigger "Alarm_Adress_4" bit 7
   13: 'Motor 4 Voltage Fault', class Errors, trigger "Alarm_Adress_4" bit 13
   14: 'Motor 4 Torque Fault', class Errors, trigger "Alarm_Adress_4" bit 14
   15: 'Motor 4 Thermal Warning', class Warnings, trigger "Alarm_Adress_4" bit 15
   16: 'Motor 5 Trip', class Errors, trigger "Alarm_Adress_5" bit 3
   17: 'Motor 5 Warning', class Warnings, trigger "Alarm_Adress_5" bit 7
   18: 'Motor 5 Voltage Fault', class Errors, trigger "Alarm_Adress_5" bit 13
   19: 'Motor 5 Torque Fault', class Errors, trigger "Alarm_Adress_5" bit 14
   20: 'Motor 5 Thermal Warning', class Warnings, trigger "Alarm_Adress_5" bit 15
   21: 'Motor 6 Trip', class Errors, trigger "Alarm_Adress_6" bit 3
   22: 'Motor 6 Warning', class Warnings, trigger "Alarm_Adress_6" bit 7
   23: 'Motor 6 Voltage Fault', class Errors, trigger "Alarm_Adress_6" bit 13
   26: 'Motor 7 Trip', class Errors, trigger "Alarm_Adress_7" bit 3
   25: 'Motor 6 Thermal Warning', class Warnings, trigger "Alarm_Adress_6" bit 15
   24: 'Motor 6 Torque Fault', class Errors, trigger "Alarm_Adress_6" bit 14
   27: 'Motor 7 Warning', class Warnings, trigger "Alarm_Adress_7" bit 7
   28: 'Motor 7 Voltage Fault', class Errors, trigger "Alarm_Adress_7" bit 13
   29: 'Motor 7 Torque Fault', class Errors, trigger "Alarm_Adress_7" bit 14
   30: 'Motor 7 Thermal Warning', class Warnings, trigger "Alarm_Adress_7" bit 15
   31: 'Motor 8 Trip', class Errors, trigger "Alarm_Adress_8" bit 3
   32: 'Motor 8 Warning', class Warnings, trigger "Alarm_Adress_8" bit 7
   33: 'Motor 8 Voltage Fault', class Errors, trigger "Alarm_Adress_8" bit 13
   34: 'Motor 8 Torque Fault', class Errors, trigger "Alarm_Adress_8" bit 14
   35: 'Motor 8 Thermal Warning', class Warnings, trigger "Alarm_Adress_8" bit 15
   36: 'Motor 9 Trip', class Errors, trigger "Alarm_Adress_9" bit 3
   37: 'Motor 9 Warning', class Warnings, trigger "Alarm_Adress_9" bit 7
   38: 'Motor 9 Voltage Fault', class Errors, trigger "Alarm_Adress_9" bit 13
   39: 'Motor 9 Torque Fault', class Errors, trigger "Alarm_Adress_9" bit 14
   40: 'Motor 9 Thermal Warning', class Warnings, trigger "Alarm_Adress_9" bit 15
   41: 'Motor 10 Trip', class Errors, trigger "Alarm_Adress_10" bit 3
   42: 'Motor 10 Warning', class Warnings, trigger "Alarm_Adress_10" bit 7
   43: 'Motor 10 Voltage Fault', class Errors, trigger "Alarm_Adress_10" bit 13
   44: 'Motor 10 Torque Fault', class Errors, trigger "Alarm_Adress_10" bit 14
   45: 'Motor 10 Thermal Warning', class Warnings, trigger "Alarm_Adress_10" bit 15
   46: 'Motor 11 Trip', class Errors, trigger "Alarm_Adress_11" bit 3
   47: 'Motor 11 Warning', class Warnings, trigger "Alarm_Adress_11" bit 7
   48: 'Motor 11 Voltage Fault', class Errors, trigger "Alarm_Adress_11" bit 13
   49: 'Motor 11 Torque Fault', class Errors, trigger "Alarm_Adress_11" bit 14
   50: 'Motor 11 Thermal Warning', class Warnings, trigger "Alarm_Adress_11" bit 15
   51: 'Motor 12 Trip', class Errors, trigger "Alarm_Adress_12" bit 3
   52: 'Motor 12 Warning', class Warnings, trigger "Alarm_Adress_12" bit 7
   53: 'Motor 12 Voltage Fault', class Errors, trigger "Alarm_Adress_12" bit 13
   54: 'Motor 12 Torque Fault', class Errors, trigger "Alarm_Adress_12" bit 14
   55: 'Motor 12 Thermal Warning', class Warnings, trigger "Alarm_Adress_12" bit 15
   56: 'Motor 13 Trip', class Errors, trigger "Alarm_Adress_13" bit 3
   57: 'Motor 13 Warning', class Warnings, trigger "Alarm_Adress_13" bit 7
   58: 'Motor 13 Voltage Fault', class Errors, trigger "Alarm_Adress_13" bit 13
   59: 'Motor 13 Torque Fault', class Errors, trigger "Alarm_Adress_13" bit 14
   60: 'Motor 13 Thermal Warning', class Warnings, trigger "Alarm_Adress_13" bit 15
   61: 'Motor 14 Trip', class Errors, trigger "Alarm_Adress_14" bit 3
   62: 'Motor 14 Warning', class Warnings, trigger "Alarm_Adress_14" bit 7
   63: 'Motor 14 Voltage Fault', class Errors, trigger "Alarm_Adress_14" bit 13
   64: 'Motor 14 Torque Fault', class Errors, trigger "Alarm_Adress_14" bit 14
   65: 'Motor 14 Thermal Warning', class Warnings, trigger "Alarm_Adress_14" bit 15
   66: 'Motor 15 Trip', class Errors, trigger "Alarm_Adress_15" bit 3
   67: 'Motor 15 Warning', class Warnings, trigger "Alarm_Adress_15" bit 7
   68: 'Motor 15 Voltage Fault', class Errors, trigger "Alarm_Adress_15" bit 13
   69: 'Motor 15 Torque Fault', class Errors, trigger "Alarm_Adress_15" bit 14
   70: 'Motor 15 Thermal Warning', class Warnings, trigger "Alarm_Adress_15" bit 15
   71: 'Motor 16 Trip', class Errors, trigger "Alarm_Adress_16" bit 3
   72: 'Motor 16 Warning', class Warnings, trigger "Alarm_Adress_16" bit 7
   73: 'Motor 16 Voltage Fault', class Errors, trigger "Alarm_Adress_16" bit 13
   74: 'Motor 16 Torque Fault', class Errors, trigger "Alarm_Adress_16" bit 14
   75: 'Motor 16 Thermal Warning', class Warnings, trigger "Alarm_Adress_16" bit 15
   76: 'Motor 17 Trip', class Errors, trigger "Alarm_Adress_17" bit 3
   77: 'Motor 17 Warning', class Warnings, trigger "Alarm_Adress_17" bit 7
   78: 'Motor 17 Voltage Fault', class Errors, trigger "Alarm_Adress_17" bit 13
   79: 'Motor 17 Torque Fault', class Errors, trigger "Alarm_Adress_17" bit 14
   80: 'Motor 17 Thermal Warning', class Warnings, trigger "Alarm_Adress_17" bit 15
   81: 'Motor 18 Trip', class Errors, trigger "Alarm_Adress_18" bit 3
   82: 'Motor 18 Warning', class Warnings, trigger "Alarm_Adress_18" bit 7
   83: 'Motor 18 Voltage Fault', class Errors, trigger "Alarm_Adress_18" bit 13
   84: 'Motor 18 Torque Fault', class Errors, trigger "Alarm_Adress_18" bit 14
   85: 'Motor 18 Thermal Warning', class Warnings, trigger "Alarm_Adress_18" bit 15
   86: 'Motor 19 Trip', class Errors, trigger "Alarm_Adress_19" bit 3
   87: 'Motor 19 Warning', class Warnings, trigger "Alarm_Adress_19" bit 7
   88: 'Motor 19 Voltage Fault', class Errors, trigger "Alarm_Adress_19" bit 13
   89: 'Motor 19 Torque Fault', class Errors, trigger "Alarm_Adress_19" bit 14
   90: 'Motor 19 Thermal Warning', class Warnings, trigger "Alarm_Adress_19" bit 15
   91: 'Motor 20 Trip', class Errors, trigger "Alarm_Adress_20" bit 3
   92: 'Motor 20 Warning', class Warnings, trigger "Alarm_Adress_20" bit 7
   93: 'Motor 20 Voltage Fault', class Errors, trigger "Alarm_Adress_20" bit 13
   94: 'Motor 20 Torque Fault', class Errors, trigger "Alarm_Adress_20" bit 14
   95: 'Motor 20 Thermal Warning', class Warnings, trigger "Alarm_Adress_20" bit 15
   96: 'Motor 21 Trip', class Errors, trigger "Alarm_Adress_21" bit 3
   97: 'Motor 21 Warning', class Warnings, trigger "Alarm_Adress_21" bit 7
   98: 'Motor 21 Voltage Fault', class Errors, trigger "Alarm_Adress_21" bit 13
   99: 'Motor 21 Torque Fault', class Errors, trigger "Alarm_Adress_21" bit 14
   100: 'Motor 21 Thermal Warning', class Warnings, trigger "Alarm_Adress_21" bit 15
   101: 'Motor 22 Trip', class Errors, trigger "Alarm_Adress_22" bit 3
   102: 'Motor 22 Warning', class Warnings, trigger "Alarm_Adress_22" bit 7
   103: 'Motor 22 Voltage Fault', class Errors, trigger "Alarm_Adress_22" bit 13
   104: 'Motor 22 Torque Fault', class Errors, trigger "Alarm_Adress_22" bit 14
   105: 'Motor 22 Thermal Warning', class Warnings, trigger "Alarm_Adress_22" bit 15
   106: 'Motor 23 Trip', class Errors, trigger "Alarm_Adress_23" bit 3
   107: 'Motor 23 Warning', class Warnings, trigger "Alarm_Adress_23" bit 7
   108: 'Motor 23 Voltage Fault', class Errors, trigger "Alarm_Adress_23" bit 13
   109: 'Motor 23 Torque Fault', class Errors, trigger "Alarm_Adress_23" bit 14
   110: 'Motor 23 Thermal Warning', class Warnings, trigger "Alarm_Adress_23" bit 15
   111: 'Profibus connection Station 2 Failure !!!', class Errors, trigger "Alarm_1" bit 9
   112: 'Profibus connection Station 3 Failure !!!', class Errors, trigger "Alarm_1" bit 10
   113: 'Profibus connection Station 4 Failure !!!', class Errors, trigger "Alarm_1" bit 11
   114: 'Profibus connection Station 5 Failure !!!', class Errors, trigger "Alarm_1" bit 12
   115: 'Profibus connection Station 6 Failure !!!', class Errors, trigger "Alarm_1" bit 13
   116: 'Profibus connection Station 7 Failure !!!', class Errors, trigger "Alarm_1" bit 14
   117: 'Profibus connection Station 8 Failure !!!', class Errors, trigger "Alarm_1" bit 15
   118: 'Profibus connection Station 9 Failure !!!', class Errors, trigger "Alarm_1" bit 0
   119: 'Profibus connection Station 10 Failure !!!', class Errors, trigger "Alarm_1" bit 1
   120: 'Profibus connection Station 11 Failure !!!', class Errors, trigger "Alarm_1" bit 2
   121: 'Profibus connection Station 12 Failure !!!', class Errors, trigger "Alarm_1" bit 3
   122: 'Profibus connection Station 13 Failure !!!', class Errors, trigger "Alarm_1" bit 4
   123: 'Profibus connection Station 14 Failure !!!', class Errors, trigger "Alarm_1" bit 5
   124: 'Profibus connection Station 15 Failure !!!', class Errors, trigger "Alarm_1" bit 6
   125: 'Profibus connection Station 16 Failure !!!', class Errors, trigger "Alarm_1" bit 7
   126: 'Profibus connection Station 17 Failure !!!', class Errors, trigger "Alarm_2" bit 8
   127: 'Profibus connection Station 18 Failure !!!', class Errors, trigger "Alarm_2" bit 9
   128: 'Profibus connection Station 19 Failure !!!', class Errors, trigger "Alarm_2" bit 10
   129: 'Profibus connection Station 20 Failure !!!', class Errors, trigger "Alarm_2" bit 11
   130: 'Profibus connection Station 21 Failure !!!', class Errors, trigger "Alarm_2" bit 12
   131: 'Profibus connection Station 22 Failure !!!', class Errors, trigger "Alarm_2" bit 13
   132: 'Profibus connection Station 23 Failure !!!', class Errors, trigger "Alarm_2" bit 14
   133: 'EMERGENCY PRESSED !!!', class Errors, trigger "Alarm_2" bit 15

text list "Mode_Syncron": 0 'Single'; 1 'Synch'

text list "Cutter_Moulder": 1 'Rotary Moulder Mode'; 2 'Rotary Cutter Mode'

text list "mde": 0 'Single'; 1 'Synchron'

